(* Logix 5000 project; controller PLC_MCC1300_75F1 vendor 1 type 14 code 166 rev 32.11; software revision 32.04; part 25 of 83 *)
(* tags used below, declared in another part *)
   CM_ConveyorStackerToLine_JS1_Sync : CM_ConveyorStackerToLine;
   GP_OB_InitializeMain : GP_OB_Initialize;
   M311 : MAC_Conveyor;
   M317 : MAC_Conveyor_Single;
   M317_ALM : MAC_Conveyor_ALM;
   M317_Data : UDT_Convoy_SL;
   M317_dTractionRecovery_M3 : DINT;
   M317_HMR : MAC_Conveyor_HMR;
   M317_HMW : MAC_Conveyor_HMW;
   M317_M1_DR_IN_MAJ : MOTION_INSTRUCTION;
   M317_M1_DR_IN_MAR : MOTION_INSTRUCTION;
   M317_M1_DR_IN_MAS : MOTION_INSTRUCTION;
   M317_M1_DR_IN_MRP : MOTION_INSTRUCTION;
   M317_M1_DR_MAFR : MOTION_INSTRUCTION;
   M317_M1_DR_MDR : MOTION_INSTRUCTION;
   M317_M1_DR_MSF : MOTION_INSTRUCTION;
   M317_M1_DR_MSO : MOTION_INSTRUCTION;
   M317_M1_DR_OUT_MAJ : MOTION_INSTRUCTION;
   M317_M1_DR_OUT_MAM : MOTION_INSTRUCTION;
   M317_M1_DR_OUT_MAR : MOTION_INSTRUCTION;
   M317_M1_DR_OUT_MAS : MOTION_INSTRUCTION;
   M317_M1_DR_OUT_MCD : MOTION_INSTRUCTION;
   M317_M1_DR_OUT_MRP : MOTION_INSTRUCTION;
   M317_M1_DR_R1 : AXIS_CIP_DRIVE;
   M317_M2_AUX_ReqSpeed_mm_min : DINT;
   M317_M2_ChangeSpeed : BOOL;
   M317_M2_DR_IN_MAJ : MOTION_INSTRUCTION;
   M317_M2_DR_IN_MAR : MOTION_INSTRUCTION;
   M317_M2_DR_IN_MAS : MOTION_INSTRUCTION;
   M317_M2_DR_IN_MRP : MOTION_INSTRUCTION;
   M317_M2_DR_MAFR : MOTION_INSTRUCTION;
   M317_M2_DR_MDR : MOTION_INSTRUCTION;
   M317_M2_DR_MSF : MOTION_INSTRUCTION;
   M317_M2_DR_MSO : MOTION_INSTRUCTION;
   M317_M2_DR_OUT_MAJ : MOTION_INSTRUCTION;
   M317_M2_DR_OUT_MAM : MOTION_INSTRUCTION;
   M317_M2_DR_OUT_MAR : MOTION_INSTRUCTION;
   M317_M2_DR_OUT_MAS : MOTION_INSTRUCTION;
   M317_M2_DR_OUT_MCD : MOTION_INSTRUCTION;
   M317_M2_DR_OUT_MRP : MOTION_INSTRUCTION;
   M317_M2_DR_R2 : AXIS_CIP_DRIVE;
   M317_M2_ReqSpeed_mm_min : DINT;
   M317_M3_AUX_ReqSpeed_mm_min : DINT;
   M317_M3_ChangeSpeed : BOOL;
   M317_M3_DR_IN_MAR : MOTION_INSTRUCTION;
   M317_M3_DR_IN_MAS : MOTION_INSTRUCTION;
   M317_M3_DR_IN_MRP : MOTION_INSTRUCTION;
   M317_M3_DR_L : AXIS_CIP_DRIVE;
   M317_M3_DR_MAFR : MOTION_INSTRUCTION;
   M317_M3_DR_MDR : MOTION_INSTRUCTION;
   M317_M3_DR_MSF : MOTION_INSTRUCTION;
   M317_M3_DR_MSO : MOTION_INSTRUCTION;
   M317_M3_DR_OUT_MAJ : MOTION_INSTRUCTION;
   M317_M3_DR_OUT_MAM : MOTION_INSTRUCTION;
   M317_M3_DR_OUT_MAR : MOTION_INSTRUCTION;
   M317_M3_DR_OUT_MRP : MOTION_INSTRUCTION;
   M317_M3_ReqSpeed_mm_min : DINT;
   M317_M3_xOSR_LatSquarFtc : BOOL;
   M317_SpaceConv_Utilities : SpaceConv_Utilities;
   M317_xOS_PosReq : BOOL;
   TMP_dDirection : DINT;
   TMP_r : REAL;
   TMP_rAcc : REAL;
   TMP_rDec : REAL;
   TMP_rSpeed : REAL;
   TMP_rTarget_M1 : REAL;
   TMP_rTarget_M2 : REAL;
   TMP_rTarget_M3 : REAL;
   TMP_xForwardCommadnForCleaningZone : BOOL;
   TMP_xPositioning_M1 : BOOL;
   TMP_xPositioning_M2 : BOOL;
   TMP_xPositioning_M3 : BOOL;
   TMP_xPowerSaving : BOOL;
   TMP_xReverse_M1 : BOOL;
   TMP_xReverse_M2 : BOOL;
   TMP_xReverse_M3 : BOOL;
   TMP_xRun_M1 : BOOL;
   TMP_xRun_M2 : BOOL;
   TMP_xRun_M3 : BOOL;
   xAlwaysOFF : BOOL;
   xDebugOFF : BOOL;
   Z402 : MAC_Zone;
   Z402_HMW : MAC_Zone_HMW;
   Z402S_INPUT_xSafetyAreaPopup : BOOL;
(* CommandLogic, continued *)

ROUTINE M317_Output   (* ladder *)
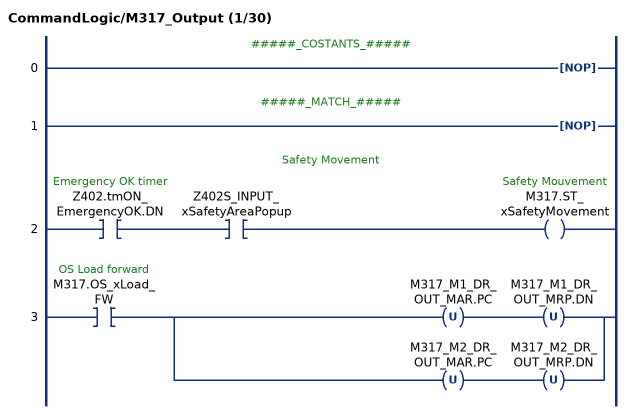
   // #####_COSTANTS_#####
   0: NOP();
   // #####_MATCH_#####
   1: NOP();
   // Safety Movement
   2: XIC(Z402.tmON_EmergencyOK.DN)XIC(Z402S_INPUT_xSafetyAreaPopup)OTE(M317.ST_xSafetyMovement);
   3: XIC(M317.OS_xLoad_FW)[OTU(M317_M1_DR_OUT_MAR.PC) OTU(M317_M1_DR_OUT_MRP.DN) ,OTU(M317_M2_DR_OUT_MAR.PC) OTU(M317_M2_DR_OUT_MRP.DN) ];
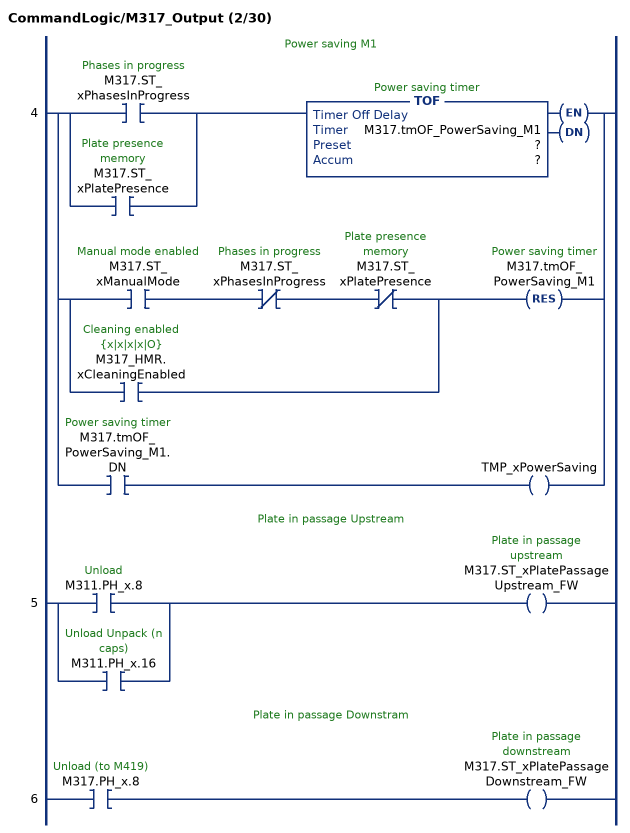
   // Power saving M1
   4: [[XIC(M317.ST_xPhasesInProgress) ,XIC(M317.ST_xPlatePresence) ] TOF(M317.tmOF_PowerSaving_M1,?,?) ,[XIC(M317.ST_xManualMode) XIO(M317.ST_xPhasesInProgress) XIO(M317.ST_xPlatePresence) ,XIC(M317_HMR.xCleaningEnabled) ] RES(M317.tmOF_PowerSaving_M1) ,XIC(M317.tmOF_PowerSaving_M1.DN) OTE(TMP_xPowerSaving) ];
   // Plate in passage Upstream
   5: [XIC(M311.PH_x.8) ,XIC(M311.PH_x.16) ]OTE(M317.ST_xPlatePassageUpstream_FW);
   // Plate in passage Downstram
   6: XIC(M317.PH_x.8)OTE(M317.ST_xPlatePassageDownstream_FW);
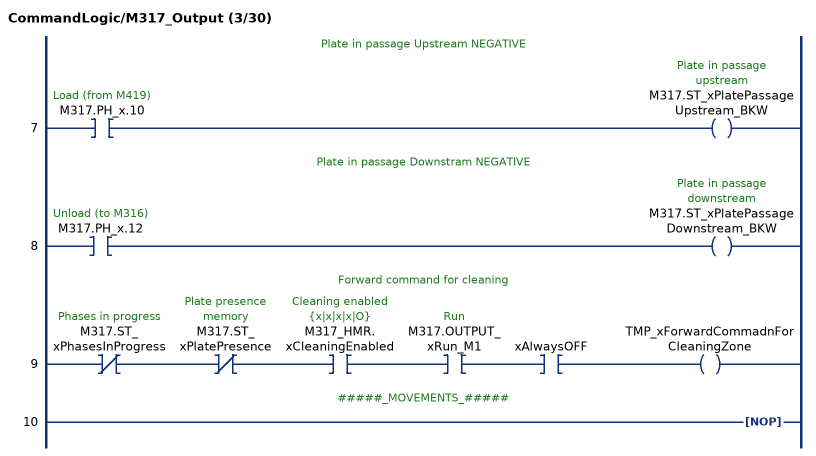
   // Plate in passage Upstream NEGATIVE
   7: XIC(M317.PH_x.10)OTE(M317.ST_xPlatePassageUpstream_BKW);
   // Plate in passage Downstram NEGATIVE
   8: XIC(M317.PH_x.12)OTE(M317.ST_xPlatePassageDownstream_BKW);
   // Forward command for cleaning
   9: XIO(M317.ST_xPhasesInProgress)XIO(M317.ST_xPlatePresence)XIC(M317_HMR.xCleaningEnabled)XIC(M317.OUTPUT_xRun_M1)XIC(xAlwaysOFF)OTE(TMP_xForwardCommadnForCleaningZone);
   // #####_MOVEMENTS_#####
   10: NOP();
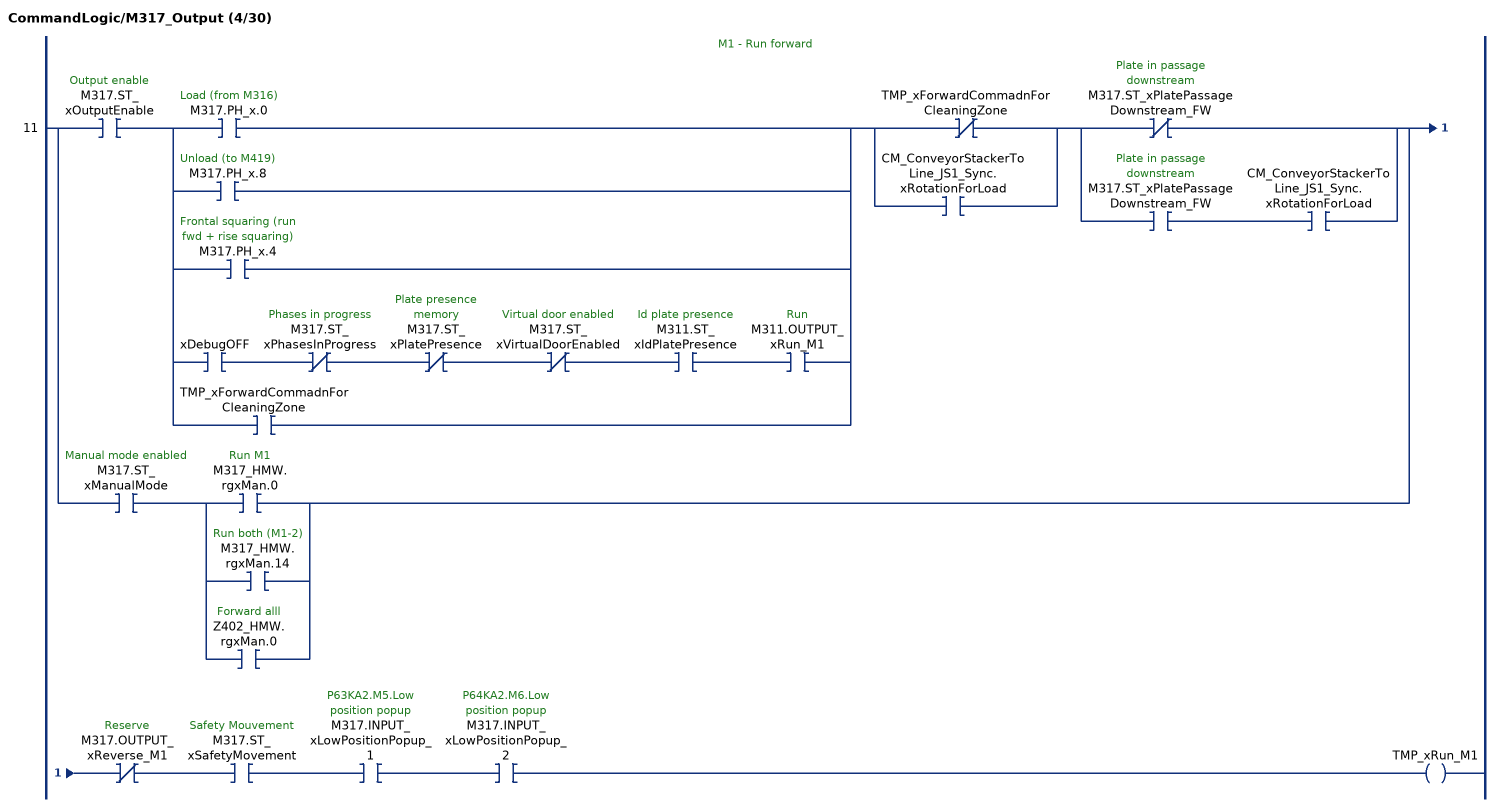
   // M1 - Run forward
   11: [XIC(M317.ST_xOutputEnable) [XIC(M317.PH_x.0) ,XIC(M317.PH_x.8) ,XIC(M317.PH_x.4) ,XIC(xDebugOFF) XIO(M317.ST_xPhasesInProgress) XIO(M317.ST_xPlatePresence) XIO(M317.ST_xVirtualDoorEnabled) XIC(M311.ST_xIdPlatePresence) XIC(M311.OUTPUT_xRun_M1) ,XIC(TMP_xForwardCommadnForCleaningZone) ] [XIO(TMP_xForwardCommadnForCleaningZone) ,XIC(CM_ConveyorStackerToLine_JS1_Sync.xRotationForLoad) ] [XIO(M317.ST_xPlatePassageDownstream_FW) ,XIC(M317.ST_xPlatePassageDownstream_FW) XIC(CM_ConveyorStackerToLine_JS1_Sync.xRotationForLoad) ] ,XIC(M317.ST_xManualMode) [XIC(M317_HMW.rgxMan.0) ,XIC(M317_HMW.rgxMan.14) ,XIC(Z402_HMW.rgxMan.0) ] ]XIO(M317.OUTPUT_xReverse_M1)XIC(M317.ST_xSafetyMovement)XIC(M317.INPUT_xLowPositionPopup_1)XIC(M317.INPUT_xLowPositionPopup_2)OTE(TMP_xRun_M1);
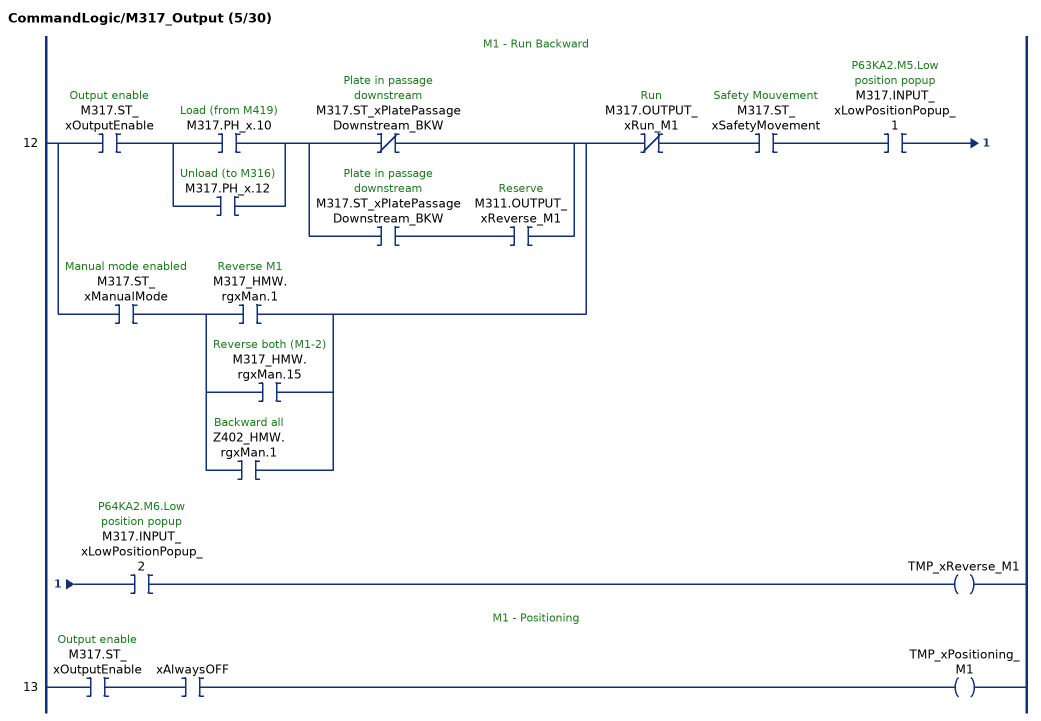
   // M1 - Run Backward
   12: [XIC(M317.ST_xOutputEnable) [XIC(M317.PH_x.10) ,XIC(M317.PH_x.12) ] [XIO(M317.ST_xPlatePassageDownstream_BKW) ,XIC(M317.ST_xPlatePassageDownstream_BKW) XIC(M311.OUTPUT_xReverse_M1) ] ,XIC(M317.ST_xManualMode) [XIC(M317_HMW.rgxMan.1) ,XIC(M317_HMW.rgxMan.15) ,XIC(Z402_HMW.rgxMan.1) ] ]XIO(M317.OUTPUT_xRun_M1)XIC(M317.ST_xSafetyMovement)XIC(M317.INPUT_xLowPositionPopup_1)XIC(M317.INPUT_xLowPositionPopup_2)OTE(TMP_xReverse_M1);
   // M1 - Positioning
   13: XIC(M317.ST_xOutputEnable)XIC(xAlwaysOFF)OTE(TMP_xPositioning_M1);
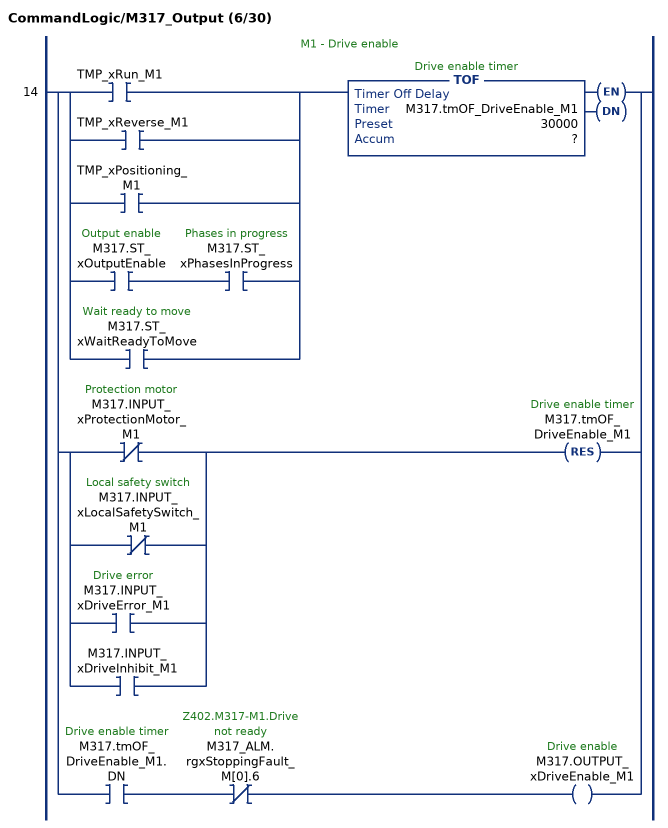
   // M1 - Drive enable
   14: [[XIC(TMP_xRun_M1) ,XIC(TMP_xReverse_M1) ,XIC(TMP_xPositioning_M1) ,XIC(M317.ST_xOutputEnable) XIC(M317.ST_xPhasesInProgress) ,XIC(M317.ST_xWaitReadyToMove) ] TOF(M317.tmOF_DriveEnable_M1,?,?) ,[XIO(M317.INPUT_xProtectionMotor_M1) ,XIO(M317.INPUT_xLocalSafetySwitch_M1) ,XIC(M317.INPUT_xDriveError_M1) ,XIC(M317.INPUT_xDriveInhibit_M1) ] RES(M317.tmOF_DriveEnable_M1) ,XIC(M317.tmOF_DriveEnable_M1.DN) XIO(M317_ALM.rgxStoppingFault_M[0].6) OTE(M317.OUTPUT_xDriveEnable_M1) ];
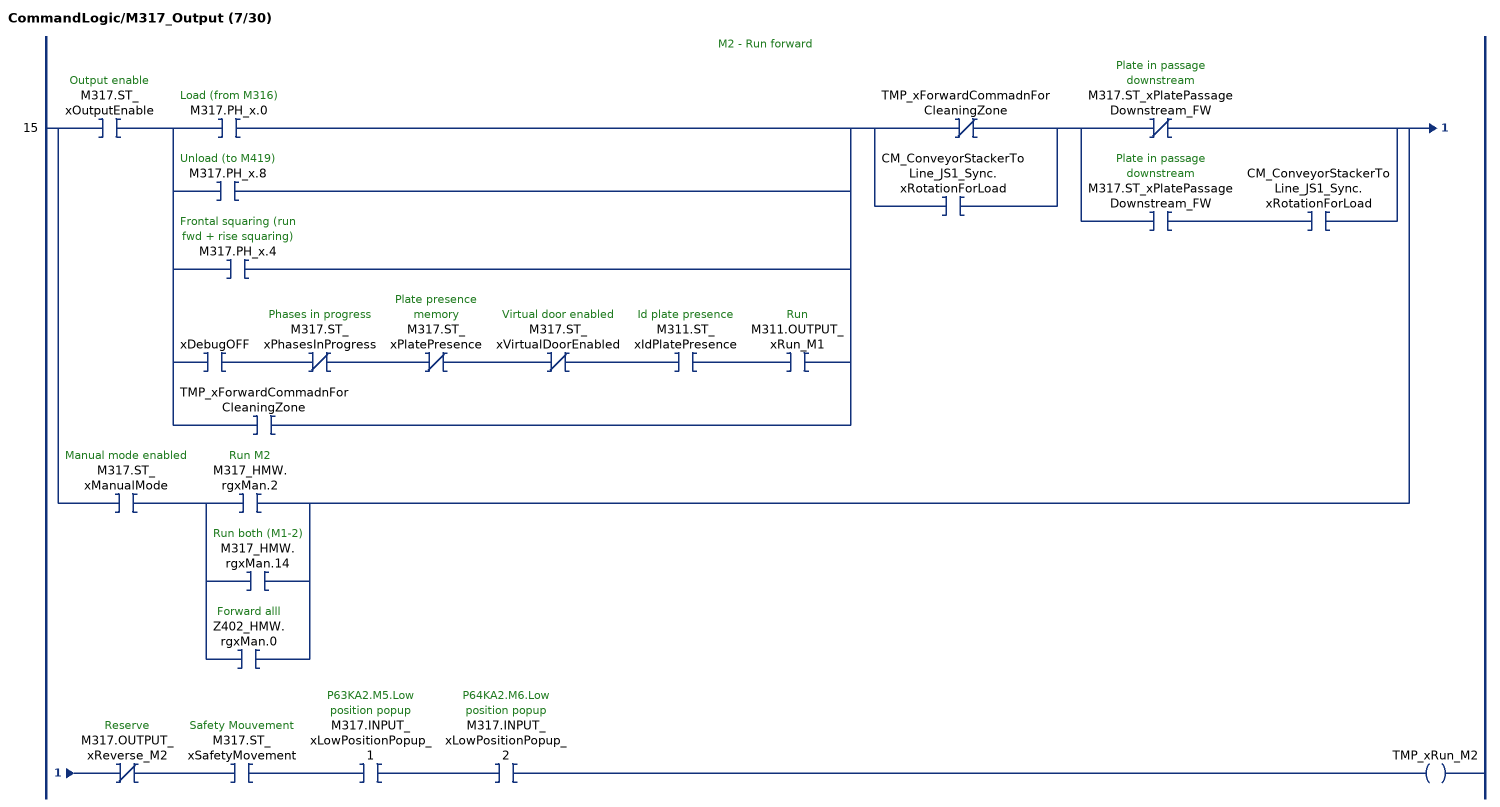
   // M2 - Run forward
   15: [XIC(M317.ST_xOutputEnable) [XIC(M317.PH_x.0) ,XIC(M317.PH_x.8) ,XIC(M317.PH_x.4) ,XIC(xDebugOFF) XIO(M317.ST_xPhasesInProgress) XIO(M317.ST_xPlatePresence) XIO(M317.ST_xVirtualDoorEnabled) XIC(M311.ST_xIdPlatePresence) XIC(M311.OUTPUT_xRun_M1) ,XIC(TMP_xForwardCommadnForCleaningZone) ] [XIO(TMP_xForwardCommadnForCleaningZone) ,XIC(CM_ConveyorStackerToLine_JS1_Sync.xRotationForLoad) ] [XIO(M317.ST_xPlatePassageDownstream_FW) ,XIC(M317.ST_xPlatePassageDownstream_FW) XIC(CM_ConveyorStackerToLine_JS1_Sync.xRotationForLoad) ] ,XIC(M317.ST_xManualMode) [XIC(M317_HMW.rgxMan.2) ,XIC(M317_HMW.rgxMan.14) ,XIC(Z402_HMW.rgxMan.0) ] ]XIO(M317.OUTPUT_xReverse_M2)XIC(M317.ST_xSafetyMovement)XIC(M317.INPUT_xLowPositionPopup_1)XIC(M317.INPUT_xLowPositionPopup_2)OTE(TMP_xRun_M2);
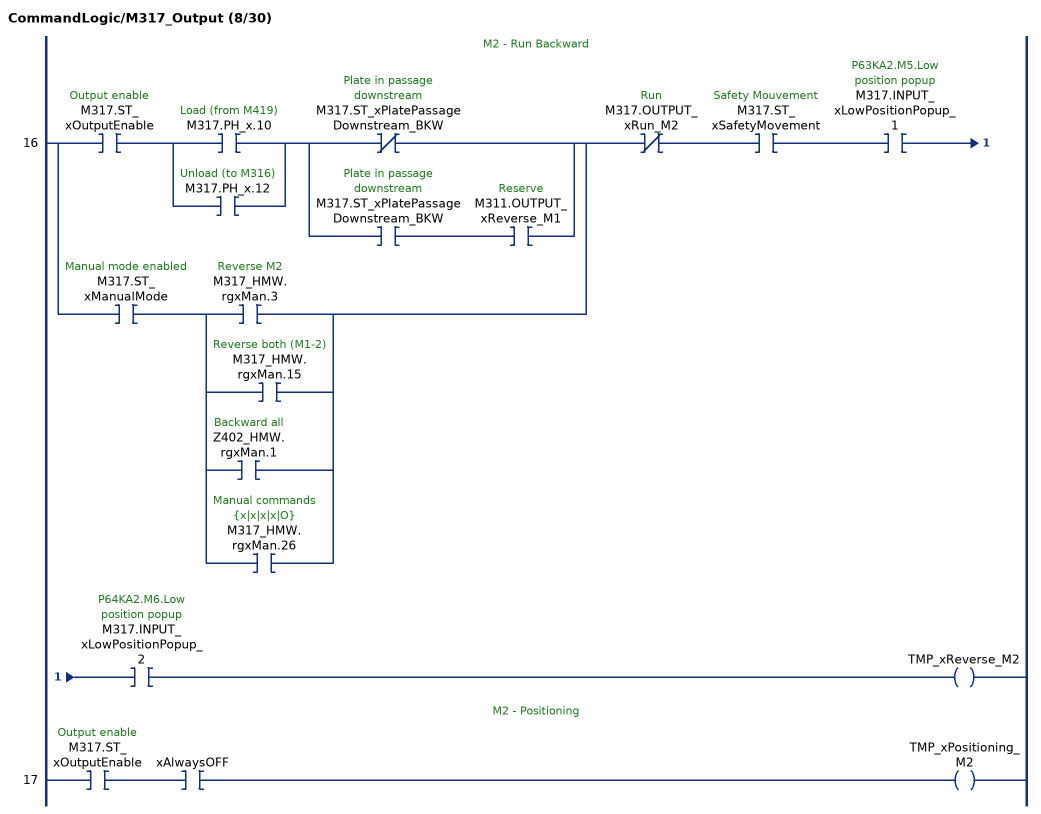
   // M2 - Run Backward
   16: [XIC(M317.ST_xOutputEnable) [XIC(M317.PH_x.10) ,XIC(M317.PH_x.12) ] [XIO(M317.ST_xPlatePassageDownstream_BKW) ,XIC(M317.ST_xPlatePassageDownstream_BKW) XIC(M311.OUTPUT_xReverse_M1) ] ,XIC(M317.ST_xManualMode) [XIC(M317_HMW.rgxMan.3) ,XIC(M317_HMW.rgxMan.15) ,XIC(Z402_HMW.rgxMan.1) ,XIC(M317_HMW.rgxMan.26) ] ]XIO(M317.OUTPUT_xRun_M2)XIC(M317.ST_xSafetyMovement)XIC(M317.INPUT_xLowPositionPopup_1)XIC(M317.INPUT_xLowPositionPopup_2)OTE(TMP_xReverse_M2);
   // M2 - Positioning
   17: XIC(M317.ST_xOutputEnable)XIC(xAlwaysOFF)OTE(TMP_xPositioning_M2);
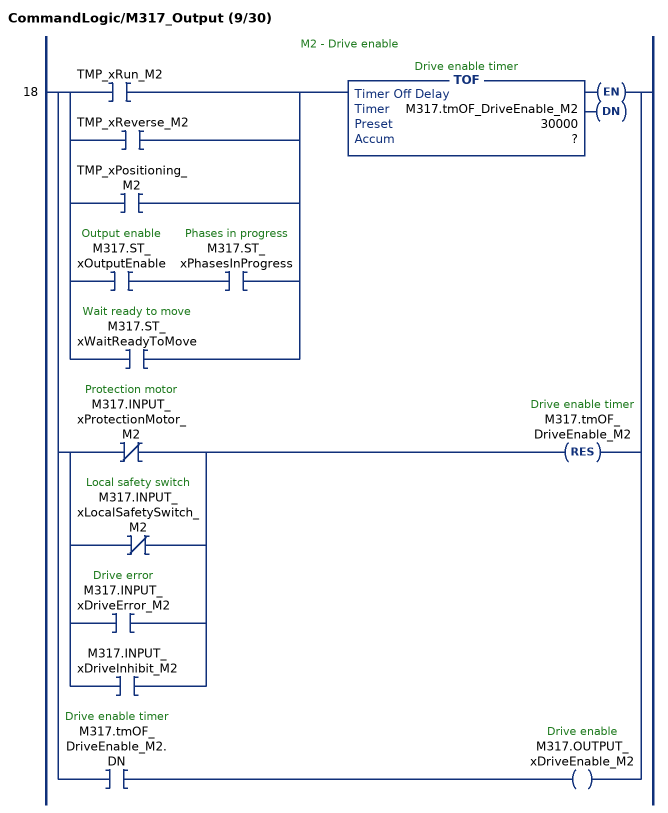
   // M2 - Drive enable
   18: [[XIC(TMP_xRun_M2) ,XIC(TMP_xReverse_M2) ,XIC(TMP_xPositioning_M2) ,XIC(M317.ST_xOutputEnable) XIC(M317.ST_xPhasesInProgress) ,XIC(M317.ST_xWaitReadyToMove) ] TOF(M317.tmOF_DriveEnable_M2,?,?) ,[XIO(M317.INPUT_xProtectionMotor_M2) ,XIO(M317.INPUT_xLocalSafetySwitch_M2) ,XIC(M317.INPUT_xDriveError_M2) ,XIC(M317.INPUT_xDriveInhibit_M2) ] RES(M317.tmOF_DriveEnable_M2) ,XIC(M317.tmOF_DriveEnable_M2.DN) OTE(M317.OUTPUT_xDriveEnable_M2) ];
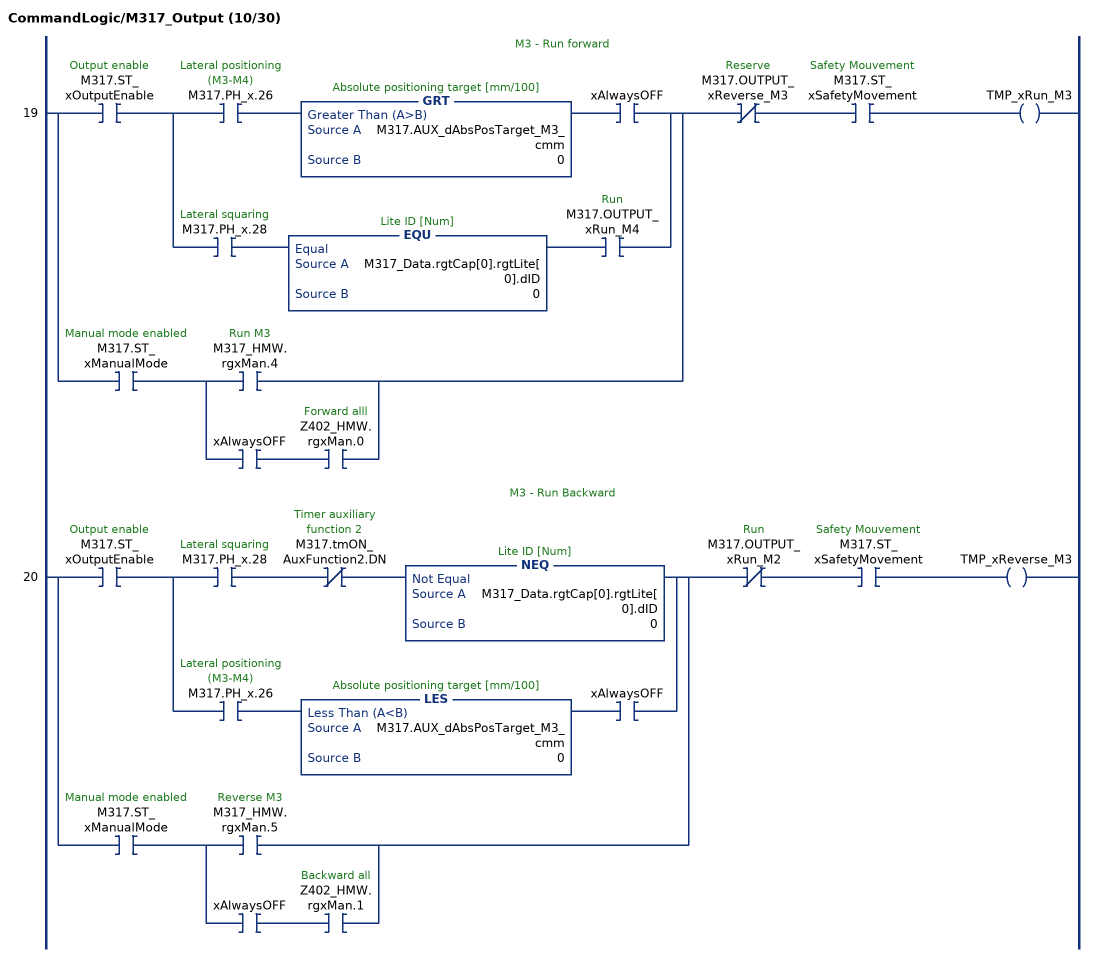
   // M3 - Run forward
   19: [XIC(M317.ST_xOutputEnable) [XIC(M317.PH_x.26) GRT(M317.AUX_dAbsPosTarget_M3_cmm,0) XIC(xAlwaysOFF) ,XIC(M317.PH_x.28) EQU(M317_Data.rgtCap[0].rgtLite[0].dID,0) XIC(M317.OUTPUT_xRun_M4) ] ,XIC(M317.ST_xManualMode) [XIC(M317_HMW.rgxMan.4) ,XIC(xAlwaysOFF) XIC(Z402_HMW.rgxMan.0) ] ]XIO(M317.OUTPUT_xReverse_M3)XIC(M317.ST_xSafetyMovement)OTE(TMP_xRun_M3);
   // M3 - Run Backward
   20: [XIC(M317.ST_xOutputEnable) [XIC(M317.PH_x.28) XIO(M317.tmON_AuxFunction2.DN) NEQ(M317_Data.rgtCap[0].rgtLite[0].dID,0) ,XIC(M317.PH_x.26) LES(M317.AUX_dAbsPosTarget_M3_cmm,0) XIC(xAlwaysOFF) ] ,XIC(M317.ST_xManualMode) [XIC(M317_HMW.rgxMan.5) ,XIC(xAlwaysOFF) XIC(Z402_HMW.rgxMan.1) ] ]XIO(M317.OUTPUT_xRun_M2)XIC(M317.ST_xSafetyMovement)OTE(TMP_xReverse_M3);
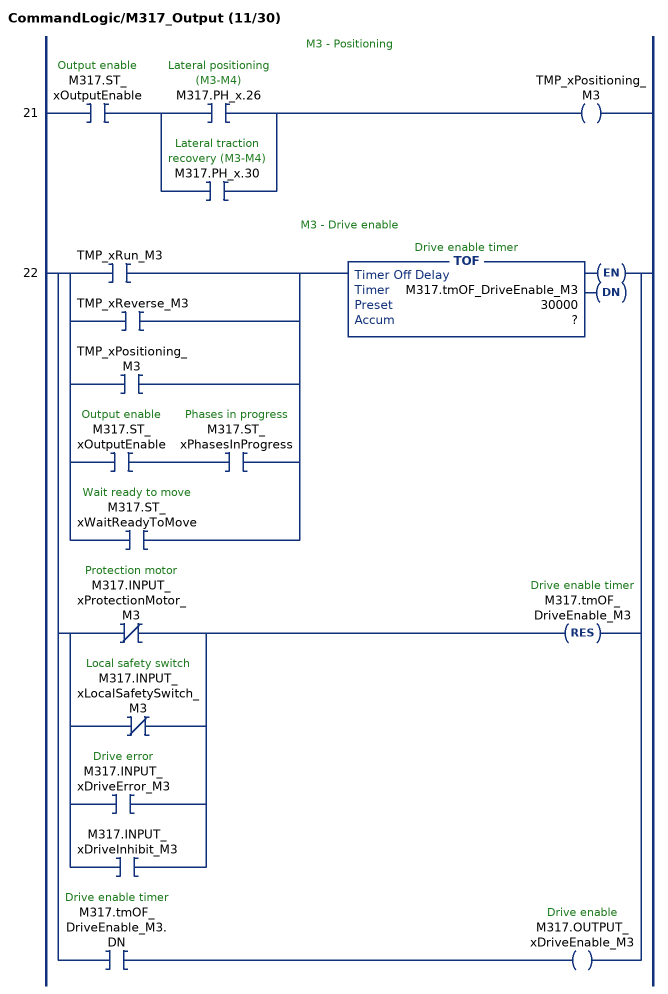
   // M3 - Positioning
   21: XIC(M317.ST_xOutputEnable)[XIC(M317.PH_x.26) ,XIC(M317.PH_x.30) ]OTE(TMP_xPositioning_M3);
   // M3 - Drive enable
   22: [[XIC(TMP_xRun_M3) ,XIC(TMP_xReverse_M3) ,XIC(TMP_xPositioning_M3) ,XIC(M317.ST_xOutputEnable) XIC(M317.ST_xPhasesInProgress) ,XIC(M317.ST_xWaitReadyToMove) ] TOF(M317.tmOF_DriveEnable_M3,?,?) ,[XIO(M317.INPUT_xProtectionMotor_M3) ,XIO(M317.INPUT_xLocalSafetySwitch_M3) ,XIC(M317.INPUT_xDriveError_M3) ,XIC(M317.INPUT_xDriveInhibit_M3) ] RES(M317.tmOF_DriveEnable_M3) ,XIC(M317.tmOF_DriveEnable_M3.DN) OTE(M317.OUTPUT_xDriveEnable_M3) ];